REGION Network 6: Fault_Mode
   // When we hit an alarm, the sequence should be aborted according to the alarm details (above in 
   // the Alarms section), and we should go into Fault mode (which is not part of our sequence).
   RUNG wire#powerrail
      Contact( "Alarm_for_E_Stop" )
      wire#w1
      Coil( "Fault_Mode" )
   END_RUNG
   RUNG wire#powerrail
      Contact( "Alarm_for_Brake_failure" )
   END_RUNG wire#w1
   RUNG wire#powerrail
      Contact( "Alarm_for_High_temp" )
   END_RUNG wire#w1
   RUNG wire#powerrail
      Contact( "Alarm_for_LOW_OIL" )
   END_RUNG wire#w1
   RUNG wire#powerrail
      Contact( "Alarm_for_Oil_High_Flow" )
   END_RUNG wire#w1
   RUNG wire#powerrail
      Contact( "Alarm_for_Over_Current" )
   END_RUNG wire#w1
   RUNG wire#powerrail
      Contact( "Alarm_for_Rotor_over_speed" )
   END_RUNG wire#w1
   // the same network as SCL:
   "Fault_Mode" := "Alarm_for_E_Stop" OR "Alarm_for_Brake_failure" OR "Alarm_for_High_temp" OR "Alarm_for_LOW_OIL" OR "Alarm_for_Oil_High_Flow" OR "Alarm_for_Over_Current" OR "Alarm_for_Rotor_over_speed";
END_REGION
END_FUNCTION_BLOCK

FUNCTION_BLOCK "HOURMETER_LAD"   // FB19, LAD
{ S7_Optimized_Access := 'TRUE' }
VERSION : 0.1
   VAR
      Min_time_down : Bool;
      Min_countdown : Bool;
      Hour_countdown : Bool;
      Day_countdown : Bool;
      Day_count_down : Bool;
      Hr_count_down : Bool;
      reset_rto : Bool;
      min_count_reset : Bool;
      hour_count_reset : Bool;
      reset_hourmeter_trigger : Bool;
      os3 : Bool;
      os2 : Bool;
      os1 : Bool;
      os4 : Bool;
      Reset_HM_Trigger : Bool;
      accum_elapsed : Time;
   END_VAR
   VAR_TEMP
      resettime : Time;
   END_VAR
   VAR_TEMP   // added for the SCL form of the ladder/FBD networks
      _w1 : Bool;
      _w2 : Bool;
      _w3 : Bool;
   END_VAR
BEGIN

REGION Network 1
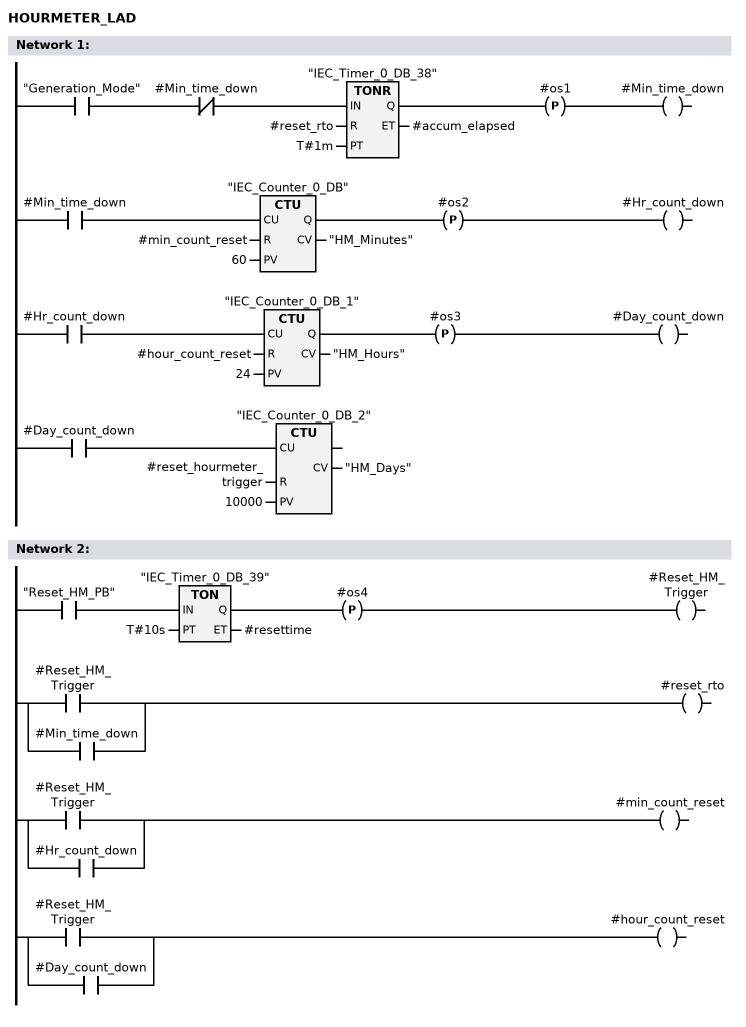
   "IEC_Timer_0_DB_38".TONR(IN := "Generation_Mode" AND NOT #Min_time_down,
                           R := #reset_rto,
                           PT := T#1m,
                           ET => #accum_elapsed);
   #_w1 := "IEC_Timer_0_DB_38".Q AND NOT #os1;   // rising edge
   #os1 := "IEC_Timer_0_DB_38".Q;
   #Min_time_down := #_w1;
   "IEC_Counter_0_DB".CTU(CU := #Min_time_down, R := #min_count_reset, PV := 60, CV => "HM_Minutes");
   #_w2 := "IEC_Counter_0_DB".Q AND NOT #os2;   // rising edge
   #os2 := "IEC_Counter_0_DB".Q;
   #Hr_count_down := #_w2;
   "IEC_Counter_0_DB_1".CTU(CU := #Hr_count_down, R := #hour_count_reset, PV := 24, CV => "HM_Hours");
   #_w3 := "IEC_Counter_0_DB_1".Q AND NOT #os3;   // rising edge
   #os3 := "IEC_Counter_0_DB_1".Q;
   #Day_count_down := #_w3;
   "IEC_Counter_0_DB_2".CTU(CU := #Day_count_down, R := #reset_hourmeter_trigger, PV := 10000, CV => "HM_Days");
END_REGION

REGION Network 2
   "IEC_Timer_0_DB_39".TON(IN := "Reset_HM_PB", PT := T#10s, ET => #resettime);
   #_w1 := "IEC_Timer_0_DB_39".Q AND NOT #os4;   // rising edge
   #os4 := "IEC_Timer_0_DB_39".Q;
   #Reset_HM_Trigger := #_w1;
   #reset_rto := #Reset_HM_Trigger OR #Min_time_down;
   #min_count_reset := #Reset_HM_Trigger OR #Hr_count_down;
   #hour_count_reset := #Reset_HM_Trigger OR #Day_count_down;
END_REGION
END_FUNCTION_BLOCK

// folder: SCL

FUNCTION_BLOCK "I/O SCL"   // FB4, SCL
{ S7_Optimized_Access := 'TRUE' }
VERSION : 0.1
BEGIN
   //Digital_Output's

   //Oil_Pump_VFD
   IF "Alarm_for_E_Stop" OR "Alarm_for_LOW_OIL" OR "VFD_HOA"=0 OR ("VFD_HOA"=2 AND NOT "OilPumpVFD_CTRL") THEN
      "OilPumpVFDen_Out" :=0;
   END_IF;

   IF "VFD_HOA"=1 OR ("VFD_HOA"=2 AND "OilPumpVFD_CTRL") AND NOT "Alarm_for_LOW_OIL" AND NOT "Alarm_for_E_Stop"  THEN
      "OilPumpVFDen_Out" := 1;
   END_IF;

   // Brake_Out
   IF "Brake_Out_HOA"=0 OR ("Brake_Out_HOA"=2 AND NOT "Brake_Out_CTRL") THEN
       "Brake_Out" := 0;
   END_IF;

   IF "Brake_Out_HOA" = 1 OR ("Brake_Out_HOA" = 2 AND "Brake_Out_CTRL") THEN
       "Brake_Out" := 1;
   END_IF;

   // Alarm Horn
   IF "Alarm_HOA" = 0 OR "Alarm_HOA" = 2 AND NOT "Alarm_CTRL" THEN
       "Alarm_horn_Q" := 0;
   END_IF;

   IF "Alarm_HOA" = 1 OR "Alarm_HOA" = 2 AND "Alarm_CTRL" THEN
       "Alarm_horn_Q" := 1;
   END_IF;

   // Station Interlock
   IF "Station_Interlock_HOA" = 0 OR "Station_Interlock_HOA" = 2 AND NOT "Station_Interlock_CTRL" THEN
       "Station_interlock" := 0;
   END_IF;

   IF "Station_Interlock_HOA" = 1 OR "Station_Interlock_HOA" = 2 AND "Station_Interlock_CTRL" THEN
       "Station_interlock" := 1;
   END_IF;




   //Analog_Output's
   "Scale_with_parameter"(input_min:=0,
                          input_signal:="Oil_pump_vfd_per",
                          input_max:=100,
                          output_max:=27648,
                          output_min:=0,
                          scaled_value=>"OilPumpVFDsp_Out");

   "Scale_with_parameter"(input_min := 0,
                          input_signal := "Baffle_per",
                          input_max := 100,
                          output_max := 27648,
                          output_min := 0,
                          scaled_value => "Baffle_Out");

    //Analog_Input's
   "Scale_with_parameter"(input_min := 0,
                          input_signal := "RPM_In",
                          input_max := 27648,
                          output_max := 200,
                          output_min := 0,
                          scaled_value => "rotor_rpm");

   "Scale_with_parameter"(input_min := 0,
                          input_signal := "OilTemp_In",
                          input_max := 27648,
                          output_max := 500,
                          output_min := 0,
                          scaled_value => "Oil_temp");

   "Scale_with_parameter"(input_min := 0,
                          input_signal := "OilFlow_In",
                          input_max := 27648,
                          output_max := 30,
                          output_min := 0,
                          scaled_value => "Oil_flow");

   "Scale_with_parameter"(input_min := 0,
                          input_signal := "Current_In",
                          input_max := 27648,
                          output_max := 700,
                          output_min := 0,
                          scaled_value => "Current_flow");

   //FULL AUTO BIT
   IF "Baffle_HOA" = 2 AND "Alarm_HOA" = 0 AND "VFD_HOA"=0 AND "Brake_Out_HOA" = 0 AND "Station_Interlock_HOA" = 0 THEN
       "FULLAUTOBIT" := 1;
   ELSE
       "FULLAUTOBIT" := 0;
   END_IF;
END_FUNCTION_BLOCK

FUNCTION_BLOCK "HOA_SCL"   // FB8, SCL
{ S7_Optimized_Access := 'TRUE' }
VERSION : 0.1
BEGIN
   //Brake ControlHOA
   IF "Brake_Out_HOA" < 0 OR "Brake_Out_HOA" > 2 THEN
       "Brake_Out_HOA" := 0;
   END_IF;

   IF "Brake_OFF_PB" AND "Brake_Out_HOA" <> 0 THEN
       "Brake_Out_HOA" := 0;
   END_IF;

   IF "Brake_HAND_PB" AND "Brake_Out_HOA" <> 1 THEN
       "Brake_Out_HOA" := 1;
   END_IF;

   IF "Brake_AUTO_PB" AND "Brake_Out_HOA" <> 2 THEN
       "Brake_Out_HOA" := 2;
   END_IF;


   //Alarm ControlHOA
   IF "Alarm_HOA" < 0 OR "Alarm_HOA" > 2 THEN
       "Alarm_HOA" := 0;
   END_IF;

   IF "Alarm_OFF_PB" AND "Alarm_HOA" <> 0 THEN
       "Alarm_HOA" := 0;
   END_IF;

   IF "Alarm_HAND_PB" AND "Alarm_HOA" <> 1 THEN
       "Alarm_HOA" := 1;
   END_IF;

   IF "Alarm_AUTO_PB" AND "Alarm_HOA" <> 2 THEN
       "Alarm_HOA" := 2;
   END_IF;

   //Station InterlockHOA
   IF "Station_Interlock_HOA" < 0 OR "Station_Interlock_HOA" > 2 THEN
       "Station_Interlock_HOA" := 0;
   END_IF;

   IF "Station_interlock_OFF_PB" AND "Station_Interlock_HOA" <> 0 THEN
       "Station_Interlock_HOA" := 0;
   END_IF;

   IF "Station_interlock_HAND_PB" AND "Station_Interlock_HOA" <> 1 THEN
       "Station_Interlock_HOA" := 1;
   END_IF;

   IF "Station_interlock_AUTO_PB" AND "Station_Interlock_HOA" <> 2 THEN
       "Station_Interlock_HOA" := 2;
   END_IF;
END_FUNCTION_BLOCK

FUNCTION_BLOCK "Alarm_SCL"   // FB12, SCL
{ S7_Optimized_Access := 'TRUE' }
VERSION : 0.1
   VAR_TEMP
      OLFD : Time;
      OLFD_AT : Bool;
      OCD : Time;
      OCD_AT : Bool;
      HOF : Time;
      HOF_AT : Bool;
      OHT : Time;
      OHT_AT : Bool;
      ROS_AT : Bool;
      ROS : Time;
      BF : Time;
      BF_AT : Bool;
      ti1 : Time;
      ti2 : Time;
      ti3 : Time;
      ti4 : Time;
      ti5 : Time;
      ti6 : Time;
      ti7 : Time;
      ti8 : Time;
   END_VAR
BEGIN
   // OIL LOW FLOW ALARM
   IF "OilPumpVFDen_Out" AND "Oil_flow" < "Oil_lowSp" AND NOT "Brake_Out" AND NOT "Alarm_for_LOW_OIL" AND NOT "Alarm_reset" THEN
       "Convert_time"(iv1 := "OilLowFlowDelaySP",
                      time1 => #OLFD);
       "IEC_Timer_0_DB_13".TON(IN := TRUE,
                               PT := #OLFD,
                               Q => #OLFD_AT,
                               ET=>#ti1);
   ELSE
       RESET_TIMER("IEC_Timer_0_DB_13");
   END_IF;

   IF #OLFD_AT THEN
       "Alarm_for_LOW_OIL" := 1;
       "Notity_for_LOW_OIL" := 1;
   END_IF;
   IF "Alarm_for_LOW_OIL" AND "Alarm_reset" THEN
       "Alarm_for_LOW_OIL" := 0;
       "Notity_for_LOW_OIL" := 0;
   END_IF;
   IF "Notity_for_LOW_OIL" AND "Notify_reset" THEN
       "Notity_for_LOW_OIL" := 0;
   END_IF;

   // OVER CURRENT ALARM
   IF "Current_flow" > "Over_currentSp" AND NOT "Alarm_for_Over_Current" AND NOT "Alarm_reset" THEN
       "Convert_time"(iv1 := "OverCurrenDelaytSP",
                      time1 => #OCD);
       "IEC_Timer_0_DB_14".TON(IN:=TRUE,
                               PT:=#OCD,
                               Q=>#OCD_AT,
                               ET=>#ti2);
   ELSE
       RESET_TIMER("IEC_Timer_0_DB_14");
   END_IF;
   IF #OCD_AT THEN
       "Alarm_for_Over_Current" := 1;
       "Notity_for_Over_Current" := 1;
   END_IF;
   IF "Alarm_for_Over_Current" AND "Alarm_reset" THEN
       "Alarm_for_Over_Current" := 0;
       "Notity_for_Over_Current" := 0;
   END_IF;
   IF "Notity_for_Over_Current" AND "Notify_reset" THEN
       "Notity_for_Over_Current" := 0;
   END_IF;

   //HIGH OIL FLOW ALARM
   IF "Oil_flow" > "Oil_highSp" AND NOT "Alarm_for_Oil_High_Flow" AND NOT "Alarm_reset" THEN
   "Convert_time"(iv1:="OilHighFlowSP",
                  time1=>#HOF);
   "IEC_Timer_0_DB_15".TON(IN:=TRUE,
                           PT:=#HOF,
                           Q=>#HOF_AT,
                           ET=>#ti3);
   ELSE
       RESET_TIMER("IEC_Timer_0_DB_15");
   END_IF;
   IF #HOF_AT THEN
       "Alarm_for_Oil_High_Flow" := 1;
       "Notity_for_Oil_High_Flow" := 1;
   END_IF;
   IF "Alarm_for_Oil_High_Flow" AND "Alarm_reset" THEN
       "Alarm_for_Oil_High_Flow" := 0;
       "Notity_for_Oil_High_Flow" := 0;
   END_IF;
   IF "Notity_for_Oil_High_Flow" AND "Notify_reset" THEN
       "Notity_for_Oil_High_Flow" := 0;
   END_IF;

   //OIL HIGH TEMP ALARM
   IF "Oil_temp" > "High_Oil_TempSp" AND NOT "Alarm_for_High_temp" AND NOT "Alarm_reset" THEN
       "Convert_time"(iv1 := "HighOilTempDelaySP",
                      time1 => #OHT);
       "IEC_Timer_0_DB_16".TON(IN:=TRUE,
                               PT:=#OHT,
                               Q=>#OHT_AT,
                               ET=>#ti4);
   ELSE
       RESET_TIMER("IEC_Timer_0_DB_16");
   END_IF;
   IF #OHT_AT THEN
       "Alarm_for_High_temp" := 1;
       "Notity_for_High_Temp" := 1;
   END_IF;
   IF "Alarm_for_High_temp" AND "Alarm_reset" THEN
       "Alarm_for_High_temp" := 0;
       "Notity_for_High_Temp" := 0;
   END_IF;
   IF "Notity_for_High_Temp" AND "Notify_reset" THEN
       "Notity_for_High_Temp" := 0;
   END_IF;

   //ROTOR SPEED ALARM
   IF "rotor_rpm" > "Rotor_Over_SpeedSp" AND NOT "Alarm_for_Rotor_over_speed" AND NOT "Alarm_reset" THEN
       "Convert_time"(iv1 := "RotorOverSpeedSP",
                      time1 => #ROS);
       "IEC_Timer_0_DB_17".TON(IN := TRUE,
                               PT := #ROS,
                               Q => #ROS_AT,
                               ET=>#ti5);
   ELSE
       RESET_TIMER("IEC_Timer_0_DB_17");
   END_IF;
   IF #ROS_AT THEN
       "Alarm_for_Rotor_over_speed" := 1;
       "Notity_for_Rotor_over_speed" := 1;
   END_IF;
   IF "Alarm_for_Rotor_over_speed" AND "Alarm_reset" THEN
       "Alarm_for_Rotor_over_speed" := 0;
       "Notity_for_Rotor_over_speed" := 0;
   END_IF;
   IF "Notity_for_Rotor_over_speed" AND "Notify_reset" THEN
       "Notity_for_Rotor_over_speed" := 0;
   END_IF;

   //BRAKE FAILURE ALARM
   IF "Brake_Out" AND "rotor_rpm" > 1 AND NOT "Alarm_for_Brake_failure" AND NOT "Alarm_reset" THEN
       "Convert_time"(iv1 := "BrakeFailureSP",
                      time1 => #BF);
       "IEC_Timer_0_DB_18".TON(IN := TRUE,
                               PT := #BF,
                               Q => #BF_AT,
                               ET=>#ti6);
   ELSE
       RESET_TIMER("IEC_Timer_0_DB_18");
   END_IF;
   IF #BF_AT THEN
       "Alarm_for_Brake_failure" := 1;
       "Notity_for_Brake_failure" := 1;
   END_IF;
   IF "Alarm_for_Brake_failure" AND "Alarm_reset" THEN
       "Alarm_for_Brake_failure" := 0;
       "Notity_for_Brake_failure" := 0;
   END_IF;
   IF "Notity_for_Brake_failure" AND "Notify_reset" THEN
       "Notity_for_Brake_failure" := 0;
   END_IF;

   //ESTOP ALARM
   IF NOT "E_Stop" AND NOT "Alarm_for_E_Stop" THEN
       "Alarm_for_E_Stop" := 1;
       "Notity_for_E_Stop" := 1;
   END_IF;
   IF "Alarm_for_E_Stop" AND "Alarm_reset" THEN
       "Alarm_for_E_Stop" := 0;
       "Notity_for_E_Stop" := 0;
   END_IF;
   IF "Notity_for_E_Stop" AND "Notify_reset" THEN
       "Notity_for_E_Stop" := 0;
   END_IF;

   //Alram Horn Ctrl
   IF "Fault_Mode" AND NOT "Alarm_CTRL" THEN
       "Alarm_CTRL" := 1;
   END_IF;
   IF "Alarm_CTRL" AND ("Alarm_reset" OR "Notify_reset") THEN
       "Alarm_CTRL" := 0;
   END_IF;
END_FUNCTION_BLOCK

FUNCTION_BLOCK "Modes_SCL"   // FB16, SCL
{ S7_Optimized_Access := 'TRUE' }
VERSION : 0.1
   VAR_TEMP
      ti1 : Time;
      Warmup_Trigger : Bool;
      t1 : Time;
      tv1 : Int;
      tv2 : Int;
      ti3 : Time;
      Stabilize_trigger : Bool;
      t2 : Time;
      ti4 : Time;
      CoolDown_trigger : Bool;
      t3 : Time;
   END_VAR
BEGIN
   // ESTOP HANDLING
   IF "Alarm_for_E_Stop" OR "Alarm_for_Brake_failure" THEN
       "Warm_Transition" := 1;
       "Stabilize_Transition" := 1;
       "Generation_Transition" := 1;
       "CoolDown_Transition" := 1;
   ELSE
       "Warm_Transition" := 0;
       "Stabilize_Transition" := 0;
       "Generation_Transition" := 0;
       "CoolDown_Transition" := 0;

       //WARM UP MODE
       IF "StartSequencePB" AND "Idle_Mode" AND "FULLAUTOBIT" THEN
           "StartSequenceBit" := 1;
       ELSE
           "StartSequenceBit" := 0;
       END_IF;
       IF "Warm_UP_Mode" THEN
           "Brake_Out_CTRL" := 0;
           "BafflePIDin" := "rotor_rpm";
           "BafflePID_SP" := "Warmup_RPM";
           "VFDsp" := "WarmUp_VFDper";
           IF "Oil_temp" > "WarmUpOilTempSp" THEN
               "Convert_time"(iv1 := "WarmUpOilDelaySp",
                              time1 => #ti1);
               "IEC_Timer_0_DB_32".TON(IN := TRUE,
                                       PT := #ti1,
                                       Q => #Warmup_Trigger,
                                       ET => #t1);
           ELSE
               RESET_TIMER("IEC_Timer_0_DB_32");
           END_IF;
           IF #Warmup_Trigger THEN
               RESET_TIMER("IEC_Timer_0_DB_32");
               "Warm_Transition" := 1;
           END_IF;
       ELSE
           "Warm_Transition" := 0;
       END_IF;
       IF "Alarm_for_Rotor_over_speed" OR "Alarm_for_High_temp" THEN
           "Warm_Transition" := 1;
       END_IF;

       //STABILIZE_MODE
       IF "Stabilize_mode" THEN
           "BafflePIDin" := "Current_flow";
           "BafflePID_SP" := "StabilizekWSP";
           #tv1 := "StabilizekWSP" - 5;
           #tv2 := "StabilizekWSP" + 5;
           IF "Current_flow" < #tv2 AND "Current_flow" > #tv1 THEN
               "Convert_time"(iv1 := "StabilizeDealySP",
                              time1 => #ti3);
               "IEC_Timer_0_DB_33".TON(IN := true,
                                       PT := #ti3,
                                       Q => #Stabilize_trigger,
                                       ET => #t2);
           ELSE
               RESET_TIMER("IEC_Timer_0_DB_33");
           END_IF;
           IF #Stabilize_trigger THEN
               RESET_TIMER("IEC_Timer_0_DB_33");
               "Stabilize_Transition" := 1;
           END_IF;
       ELSE
           "Stabilize_Transition" := 0;
       END_IF;
       IF "Alarm_for_Rotor_over_speed" OR "Alarm_for_High_temp" THEN
           "Stabilize_Transition" := 1;
       END_IF;

       // GENERATION MODE
       IF "Generation_Mode" THEN
           "Station_Interlock_CTRL" := 1;
           IF "System_Stop_PB" THEN
               "Generation_Transition" := 1;
           END_IF;
       ELSE
           "Generation_Transition" := 0;
       END_IF;

       IF "Alarm_for_Over_Current" OR "Alarm_for_Rotor_over_speed" OR "Alarm_for_High_temp" THEN
           "Generation_Transition" := 1;
       END_IF;
   END_IF;

           //COOLDOWN MODE
       IF "CoolDown_Mode" THEN
           "Station_Interlock_CTRL" := 0;
           "BafflePIDin" := "rotor_rpm";
           "BafflePID_SP" := "CoolDown_RPM";
           IF "Oil_temp" < "CoolDownOilTempSp" THEN
               "Convert_time"(iv1 := "CoolDownlDelaySp",
                              time1 => #ti4);
               "IEC_Timer_0_DB_34".TON(IN := true,
                                       PT := #ti4,
                                       Q => #CoolDown_trigger,
                                       ET => #t3);
           ELSE
               RESET_TIMER("IEC_Timer_0_DB_34");
           END_IF;
           IF #CoolDown_trigger THEN
               RESET_TIMER("IEC_Timer_0_DB_34");
               "CoolDown_Transition" := 1;
           END_IF;
       ELSE
           "CoolDown_Transition" := 0;
       END_IF;


       // FAULT MODE
       IF "Alarm_for_Brake_failure" OR "Alarm_for_E_Stop" OR "Alarm_for_High_temp" OR "Alarm_for_LOW_OIL" OR "Alarm_for_Oil_High_Flow" OR "Alarm_for_Over_Current" OR "Alarm_for_Rotor_over_speed" THEN
           "Fault_Mode" := 1;
       ELSE
           "Fault_Mode" := 0;
       END_IF;


   //IDLE MODE
   IF "Idle_Mode" THEN
       "Brake_Out_CTRL" := 1;
       "Baffle_Ctrl" := 0;
       "OilPumpVFD_CTRL" := 0;
       "Station_Interlock_CTRL" := 0;
   END_IF;
END_FUNCTION_BLOCK

FUNCTION_BLOCK "HOURMETER_SCL"   // FB21, SCL
{ S7_Optimized_Access := 'TRUE' }
VERSION : 0.1
   VAR
      Min_time_down : Bool;
      Min_countdown : Bool;
      Hour_countdown : Bool;
      Day_countdown : Bool;
      Day_count_down : Bool;
      Hr_count_down : Bool;
      reset_rto : Bool;
      min_count_reset : Bool;
      hour_count_reset : Bool;
      reset_hourmeter_trigger : Bool;
      os3 : Bool;
      os2 : Bool;
      os1 : Bool;
      os4 : Bool;
      Reset_HM_Trigger : Bool;
      accum_elapsed : Time;
   END_VAR
   VAR_TEMP
      resettime : Time;
   END_VAR
BEGIN
   IF "Generation_Mode" AND NOT #Min_time_down THEN
      "IEC_Timer_0_DB_42".TONR(IN := TRUE,
                                R := #reset_rto,
                                PT := t#60s,
                                Q => #Min_time_down,
                                ET => #accum_elapsed);
                            END_IF;

   IF #Min_time_down THEN
       RESET_TIMER("IEC_Timer_0_DB_42");
   END_IF;

   IF #Min_time_down THEN
       "IEC_Counter_0_DB_6".CTU(CU := #Min_time_down,
                                R := #min_count_reset,
                                PV := 60,
                                Q => #Hr_count_down,
                                CV => "HM_Minutes");
   END_IF;

   IF #Hr_count_down THEN
       "IEC_Counter_0_DB_7".CTU(CU := #Hr_count_down,
                                R := #hour_count_reset,
                                PV := 24,
                                Q => #Day_count_down,
                                CV => "HM_Hours");
   END_IF;

   IF #Day_count_down THEN

       "IEC_Counter_0_DB_8".CTU(CU := #Day_count_down,
                                R := #reset_hourmeter_trigger,
                                PV := 1000,
                                CV => "HM_Days");
   END_IF;

   IF "Reset_HM_PB" THEN
       "IEC_Timer_0_DB_43".TON(IN := TRUE,
                               PT := T#10s,
                               Q => #Reset_HM_Trigger,
                               ET => #resettime);
   ELSE
       RESET_TIMER("IEC_Timer_0_DB_43");
   END_IF;

   IF #Reset_HM_Trigger OR #Min_time_down THEN
       #reset_rto := 1;
   ELSE
       #reset_rto := 0;
   END_IF;

   IF #Reset_HM_Trigger OR #Hr_count_down THEN
       #min_count_reset := 1;
   ELSE
       #min_count_reset := 0;
   END_IF;

   IF #Reset_HM_Trigger OR #Day_count_down THEN
       #hour_count_reset := 1;
   ELSE
       #hour_count_reset := 0;
   END_IF;
END_FUNCTION_BLOCK

// folder: STL

FUNCTION_BLOCK "I/O STL"   // FB5, STL
{ S7_Optimized_Access := 'TRUE' }
VERSION : 0.1
BEGIN

REGION Network 1
   //Digital_Output's

   OilPumpVFD:A     "Alarm_for_LOW_OIL";
         JC    ResetOilPumpVFD;
         CLR;
         A     "Alarm_for_E_Stop";
         JC    ResetOilPumpVFD;
         L     "VFD_HOA";
         L     0;
         ==I;
         JC    ResetOilPumpVFD;
         CLR;
         L     "VFD_HOA";
         L     1;
         ==I;
         JC    SetoilPumpVFD;
         CLR;
         L     "VFD_HOA";
         L     2;
         ==I;
         JC    SetoilPumpVFD;
   AutoOilPumpVFD:A     "OilPumpVFD_CTRL";
         JC    SetoilPumpVFD;
         JU    ResetOilPumpVFD;

   SetoilPumpVFD:AN    "Alarm_for_LOW_OIL";
         AN    "Alarm_for_E_Stop";
         S     "OilPumpVFDen_Out";
         JU    Brake_Out;
   ResetOilPumpVFD:R     "OilPumpVFDen_Out";
         JU    Brake_Out;


   Brake_Out:L     "Brake_Out_HOA";
         L     0;
         ==I;
         JC    ResetBrake_Out;
         CLR;
         L     "Brake_Out_HOA";
         L     1;
         ==I;
         JC    SetBrake_Out;
         CLR;
         L     "Brake_Out_HOA";
         L     2;
         ==I;
         JC    SetBrake_Out;
   AutoBrake_Out:A     "Brake_Out_CTRL";
         JC    SetBrake_Out;
         JU    ResetBrake_Out;

   SetBrake_Out:S     "Brake_Out";
         JU    Alarm_horn;
   ResetBrake_Out:R     "Brake_Out";
         JU    Alarm_horn;


   Alarm_horn:L     "Alarm_HOA";
         L     0;
         ==I;
         JC    ResetAlarm_Horn;
         CLR;
         L     "Alarm_HOA";
         L     1;
         ==I;
         JC    SetAlarm_Horn;
         CLR;
         L     "Alarm_HOA";
         L     2;
         ==I;
         JC    SetAlarm_Horn;
   AutoAlarm_Horn:A     "Alarm_CTRL";
         JC    SetAlarm_Horn;
         JU    ResetAlarm_Horn;

   SetAlarm_Horn:S     "Alarm_horn_Q";
         JU    Station_Interlock;
   ResetAlarm_Horn:R     "Alarm_horn_Q";
         JU    Station_Interlock;


   Station_Interlock:A     "Alarm_for_E_Stop";
         JC    ResetStation_interlock;
         L     "Station_Interlock_HOA";
         L     0;
         ==I;
         JC    ResetStation_interlock;
         CLR;
         L     "Station_Interlock_HOA";
         L     1;
         ==I;
         JC    SetStation_interlock;
         CLR;
         L     "Station_Interlock_HOA";
         L     2;
         ==I;
         JC    SetStation_interlock;
   AutoStation_interlock:A     "Station_Interlock_CTRL";
         JC    SetStation_interlock;
         JU    ResetStation_interlock;

   SetStation_interlock:S     "Station_interlock";
         AN    "Alarm_for_E_Stop";
         JU    Analog_Output;
   ResetStation_interlock:R     "Station_interlock";
         JU    Analog_Output;



   //Analog_Output's

   Analog_Output:CALL  "Scale_with_parameter"
         ( input_min    := 0,
           input_signal := "Oil_pump_vfd_per",
           input_max    := 100,
           output_max   := 27648,
           output_min   := 0,
           scaled_value := "OilPumpVFDsp_Out"
         );

         CALL  "Scale_with_parameter"
         ( input_min    := 0,
           input_signal := "Baffle_per",
           input_max    := 100,
           output_max   := 27648,
           output_min   := 0,
           scaled_value := "Baffle_Out"
         );

   //Analog_Input's
   Analog_Input:CALL  "Scale_with_parameter"
         ( input_min    := 0,
           input_signal := "OilTemp_In",
           input_max    := 27648,
           output_max   := 500,
           output_min   := 0,
           scaled_value := "Oil_temp"
         );

         CALL  "Scale_with_parameter"
         ( input_min    := 0,
           input_signal := "OilFlow_In",
           input_max    := 27648,
           output_max   := 30,
           output_min   := 0,
           scaled_value := "Oil_flow"
         );

         CALL  "Scale_with_parameter"
         ( input_min    := 0,
           input_signal := "RPM_In",
           input_max    := 27648,
           output_max   := 200,
           output_min   := 0,
           scaled_value := "rotor_rpm"
         );

         CALL  "Scale_with_parameter"
         ( input_min    := 0,
           input_signal := "Current_In",
           input_max    := 27648,
           output_max   := 700,
           output_min   := 0,
           scaled_value := "Current_flow"
         );

   //FULL AUTO BIT
         CLR;
         L     "Baffle_HOA";
         L     2;
         ==I;
         NOT;
         JC    ResetFullAuto;
         CLR;
         L     "VFD_HOA";
         L     2;
         ==I;
         NOT;
         JC    ResetFullAuto;
         CLR;
         L     "Alarm_HOA";
         L     2;
         ==I;
         NOT;
         JC    ResetFullAuto;
         CLR;
         L     "Brake_Out_HOA";
         L     2;
         ==I;
         NOT;
         JC    ResetFullAuto;
         CLR;
         L     "Station_Interlock_HOA";
         L     2;
         ==I;
         NOT;
         JC    ResetFullAuto;
         CLR;
         SET;
         S     "FULLAUTOBIT";
         JU    endofline;

   ResetFullAuto:SET;
         NOT;
         R     "FULLAUTOBIT";
         JU    endofline;


   endofline:BE;
END_REGION
END_FUNCTION_BLOCK

FUNCTION_BLOCK "HOA_STL"   // FB9, STL
{ S7_Optimized_Access := 'TRUE' }
VERSION : 0.1
   VAR
      OS1 : Bool;
      OS2 : Bool;
      OS3 : Bool;
      OS4 : Bool;
      OS5 : Bool;
      OS6 : Bool;
      OS7 : Bool;
      OS8 : Bool;
      OS9 : Bool;
      OS10 : Bool;
      OS11 : Bool;
      OS12 : Bool;
   END_VAR
BEGIN

REGION Network 1
         L     "Brake_Out_HOA";
         L     0;
         <I;
         JC    SetBrakeoutHOAZero;
         CLR;
         L     "Brake_Out_HOA";
         L     2;
         >I;
         JC    SetBrakeoutHOAZero;
         CLR;
         A     "Brake_OFF_PB";
         FP    #OS4;
         JC    SetBrakeoutHOAZero;
         CLR;
         A     "Brake_HAND_PB";
         FP    #OS5;
         JC    SetBrakeoutHOAOne;
         CLR;
         A     "Brake_AUTO_PB";
         FP    #OS6;
         JC    SetBrakeoutHOATwo;
         JU    Alarm_Horn;

   SetBrakeoutHOAZero:L     0;
         T     "Brake_Out_HOA";
         JU    Alarm_Horn;
   SetBrakeoutHOAOne:L     1;
         T     "Brake_Out_HOA";
         JU    Alarm_Horn;
   SetBrakeoutHOATwo:L     2;
         T     "Brake_Out_HOA";
         JU    Alarm_Horn;


   Alarm_Horn:L     "Alarm_HOA";
         L     0;
         <I;
         JC    SetAlarmHOAZero;
         CLR;
         L     "Alarm_HOA";
         L     2;
         >I;
         JC    SetAlarmHOAZero;
         CLR;
         A     "Alarm_OFF_PB";
         FP    #OS7;
         JC    SetAlarmHOAZero;
         CLR;
         A     "Alarm_HAND_PB";
         FP    #OS8;
         JC    SetAlarmHOAOne;
         CLR;
         A     "Alarm_AUTO_PB";
         FP    #OS9;
         JC    SetAlarmHOATwo;
         JU    Station_Interlock;

   SetAlarmHOAZero:L     0;
         T     "Alarm_HOA";
         JU    Station_Interlock;
   SetAlarmHOAOne:L     1;
         T     "Alarm_HOA";
         JU    Station_Interlock;
   SetAlarmHOATwo:L     2;
         T     "Alarm_HOA";
         JU    Station_Interlock;


   Station_Interlock:L     "Station_Interlock_HOA";
         L     0;
         <I;
         JC    SetStationInterlockHOAZero;
         CLR;
         L     "Station_Interlock_HOA";
         L     2;
         >I;
         JC    SetStationInterlockHOAZero;
         CLR;
         A     "Station_interlock_OFF_PB";
         FP    #OS10;
         JC    SetStationInterlockHOAZero;
         CLR;
         A     "Station_interlock_HAND_PB";
         FP    #OS11;
         JC    SetStationInterlockHOAOne;
         CLR;
         A     "Station_interlock_AUTO_PB";
         FP    #OS12;
         JC    SetStationInterlockHOATwo;
         JU    Endofline;

   SetStationInterlockHOAZero:L     0;
         T     "Station_Interlock_HOA";
         BE;
   SetStationInterlockHOAOne:L     1;
         T     "Station_Interlock_HOA";
         BE;
   SetStationInterlockHOATwo:L     2;
         T     "Station_Interlock_HOA";
         BE;
   Endofline:BE;
END_REGION
END_FUNCTION_BLOCK

FUNCTION_BLOCK "Alarm_STL"   // FB13, STL
{ S7_Optimized_Access := 'TRUE' }
VERSION : 0.1
   VAR
      os1 : Bool;
      os2 : Bool;
      os3 : Bool;
      os4 : Bool;
      os5 : Bool;
      os6 : Bool;
      os7 : Bool;
      os8 : Bool;
      os9 : Bool;
      os10 : Bool;
      os11 : Bool;
      os12 : Bool;
      os13 : Bool;
      os14 : Bool;
      os15 : Bool;
      os16 : Bool;
      os17 : Bool;
   END_VAR
   VAR_TEMP
      TI_1 : Time;
      TI_2 : Time;
      TI_3 : Time;
      TI_4 : Time;
      TI_5 : Time;
      TI_6 : Time;
      T1 : Time;
      T2 : Time;
      T3 : Time;
      T4 : Time;
      T5 : Time;
      T6 : Time;
      OLFD_AT : Bool;
      OCD_AT : Bool;
      OFH_AT : Bool;
      HOT_AT : Bool;
      ROS_AT : Bool;
      BF_AT : Bool;
   END_VAR
BEGIN

REGION Network 1
   //OIL LOW FLOW ALARM
   Oil_Low_Flow:A     "Alarm_reset";
         FP    #os1;
         JC    ResetOfAlaram;
         CLR;
         A     "Notify_reset";
         FP    #os2;
         JC    ResetOfNotify;
         CLR;
         L     "Oil_flow";
         L     "Oil_lowSp";
         <I;
         A     "OilPumpVFDen_Out";
         AN    "Brake_Out";
         JC    TIMERFOROLF;
         JU    Over_current;

   TIMERFOROLF:CALL  "Convert_time"
         ( iv1   := "OilLowFlowDelaySP",
           time1 := #TI_1
         );
         CALL  TON, "IEC_Timer_0_DB_19"
         ( IN := true,
           PT := #TI_1,
           Q  := #OLFD_AT,
           ET := #T1
         );
         A     #OLFD_AT;
         JC    SetOfAlarm;
         JU    Over_current;

   SetOfAlarm:SET;
         S     "Alarm_for_LOW_OIL";
         S     "Notity_for_LOW_OIL";
         JU    Over_current;

   ResetOfAlaram:R     "Alarm_for_LOW_OIL";
         R     "Notity_for_LOW_OIL";
         CALL  RESET_TIMER
         ( "TIMER" := "IEC_Timer_0_DB_19"
         );
         JU    Over_current;

   ResetOfNotify:R     "Notity_for_LOW_OIL";
         JU    Over_current;


   //OVER CURRENT ALARM
   Over_current:A     "Alarm_reset";
         FP    #os3;
         JC    ResetOfAlaramOC;
         CLR;
         A     "Notify_reset";
         FP    #os4;
         JC    ResetOfNotifyOC;
         CLR;
         L     "Current_flow";
         L     "Over_currentSp";
         >I;
         JC    TIMERFOROC;
         JU    Oil_Flow_high;

   TIMERFOROC:CALL  "Convert_time"
         ( iv1   := "OverCurrenDelaytSP",
           time1 := #TI_2
         );
         CALL  TON , "IEC_Timer_0_DB_20"
         ( IN := true,
           PT := #TI_2,
           Q  := #OCD_AT,
           ET := #T2
         );
         A     #OCD_AT;
         JC    SetOfAlarmOC;
         JU    Oil_Flow_high;

   SetOfAlarmOC:SET;
         S     "Alarm_for_Over_Current";
         S     "Notity_for_Over_Current";
         JU    Oil_Flow_high;

   ResetOfAlaramOC:R     "Alarm_for_Over_Current";
         R     "Notity_for_Over_Current";
         CALL  RESET_TIMER
         ( "TIMER" := "IEC_Timer_0_DB_20"
         );
         JU    Oil_Flow_high;

   ResetOfNotifyOC:R     "Notity_for_Over_Current";
         JU    Oil_Flow_high;


   //OIL FLOW HIGH ALARM
   Oil_Flow_high:A     "Alarm_reset";
         FP    #os5;
         JC    ResetOfAlaramOFH;
         CLR;
         A     "Notify_reset";
         FP    #os6;
         JC    ResetOfNotifyOFH;
         CLR;
         L     "Oil_flow";
         L     "Oil_highSp";
         >I;
         JC    TIMERFOROFH;
         JU    High_Oil_Temp;


   TIMERFOROFH:CALL  "Convert_time"
         ( iv1   := "OilHighFlowSP",
           time1 := #TI_3
         );
         CALL  TON , "IEC_Timer_0_DB_21"
         ( IN := true,
           PT := #TI_3,
           Q  := #OFH_AT,
           ET := #T3
         );
         A     #OFH_AT;
         JC    SetOfAlarmOFH;
         JU    High_Oil_Temp;

   SetOfAlarmOFH:SET;
         S     "Alarm_for_Oil_High_Flow";
         S     "Notity_for_Oil_High_Flow";
         JU    High_Oil_Temp;

   ResetOfAlaramOFH:R     "Alarm_for_Oil_High_Flow";
         R     "Notity_for_Oil_High_Flow";
         CALL  RESET_TIMER
         ( "TIMER" := "IEC_Timer_0_DB_21"
         );
         JU    High_Oil_Temp;

   ResetOfNotifyOFH:R     "Notity_for_Oil_High_Flow";
         JU    High_Oil_Temp;


   //HIGH OIL TEMP ALARM
   High_Oil_Temp:A     "Alarm_reset";
         FP    #os7;
         JC    ResetOfAlaramHOT;
         CLR;
         A     "Notify_reset";
         FP    #os8;
         JC    ResetOfNotifyHOT;
         CLR;
         L     "Oil_temp";
         L     "High_Oil_TempSp";
         >I;
         JC    TIMERFORHOT;
         JU    Rotor_Over_Speed;

   TIMERFORHOT:CALL  "Convert_time"
         ( iv1   := "HighOilTempDelaySP",
           time1 := #TI_4
         );
         CALL  TON , "IEC_Timer_0_DB_22"
         ( IN := true,
           PT := #TI_4,
           Q  := #HOT_AT,
           ET := #T4
         );
         A     #HOT_AT;
         JC    SetOfAlarmHOT;
         JU    Rotor_Over_Speed;

   SetOfAlarmHOT:SET;
         S     "Alarm_for_High_temp";
         S     "Notity_for_High_Temp";
         JU    Rotor_Over_Speed;

   ResetOfAlaramHOT:R     "Alarm_for_High_temp";
         R     "Notity_for_High_Temp";
         CALL  RESET_TIMER
         ( "TIMER" := "IEC_Timer_0_DB_22"
         );
         JU    Rotor_Over_Speed;

   ResetOfNotifyHOT:R     "Notity_for_High_Temp";
         JU    Rotor_Over_Speed;


   //ROTOR OVER SPEED ALARM
   Rotor_Over_Speed:A     "Alarm_reset";
         FP    #os9;
         JC    ResetOfAlaramROS;
         CLR;
         A     "Notify_reset";
         FP    #os10;
         JC    ResetOfNotifyROS;
         CLR;
         L     "rotor_rpm";
         L     "Rotor_Over_SpeedSp";
         >I;
         JC    TIMERFORROS;
         JU    Brake_Failure;

   TIMERFORROS:CALL  "Convert_time"
         ( iv1   := "RotorOverSpeedSP",
           time1 := #TI_5
         );
         CALL  TON , "IEC_Timer_0_DB_23"
         ( IN := true,
           PT := #TI_5,
           Q  := #ROS_AT,
           ET := #T5
         );
         A     #ROS_AT;
         JC    SetOfAlarmROS;
         JU    Brake_Failure;

   SetOfAlarmROS:SET;
         S     "Alarm_for_Rotor_over_speed";
         S     "Notity_for_Rotor_over_speed";
         JU    Brake_Failure;

   ResetOfAlaramROS:R     "Alarm_for_Rotor_over_speed";
         R     "Notity_for_Rotor_over_speed";
         CALL  RESET_TIMER
         ( "TIMER" := "IEC_Timer_0_DB_23"
         );
         JU    Brake_Failure;